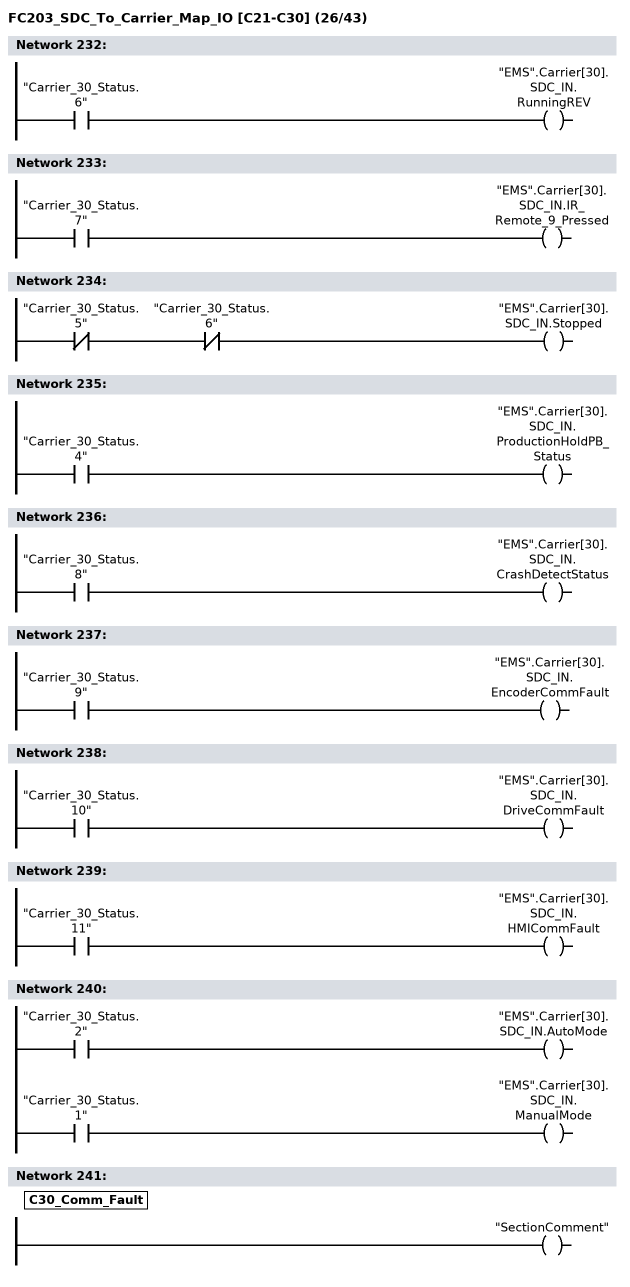
   RUNG wire#powerrail
      Contact( "Carrier_30_Status.6" )
      Coil( "EMS".Carrier[30].SDC_IN.RunningREV )
   END_RUNG
   // the same network as SCL:
   "EMS".Carrier[30].SDC_IN.RunningREV := "Carrier_30_Status.6";
END_REGION

REGION Network 233
   RUNG wire#powerrail
      Contact( "Carrier_30_Status.7" )
      Coil( "EMS".Carrier[30].SDC_IN.IR_Remote_9_Pressed )
   END_RUNG
   // the same network as SCL:
   "EMS".Carrier[30].SDC_IN.IR_Remote_9_Pressed := "Carrier_30_Status.7";
END_REGION

REGION Network 234
   RUNG wire#powerrail
      I_Contact( "Carrier_30_Status.5" )
      I_Contact( "Carrier_30_Status.6" )
      Coil( "EMS".Carrier[30].SDC_IN.Stopped )
   END_RUNG
   // the same network as SCL:
   "EMS".Carrier[30].SDC_IN.Stopped := NOT "Carrier_30_Status.5" AND NOT "Carrier_30_Status.6";
END_REGION

REGION Network 235
   RUNG wire#powerrail
      Contact( "Carrier_30_Status.4" )
      Coil( "EMS".Carrier[30].SDC_IN.ProductionHoldPB_Status )
   END_RUNG
   // the same network as SCL:
   "EMS".Carrier[30].SDC_IN.ProductionHoldPB_Status := "Carrier_30_Status.4";
END_REGION

REGION Network 236
   RUNG wire#powerrail
      Contact( "Carrier_30_Status.8" )
      Coil( "EMS".Carrier[30].SDC_IN.CrashDetectStatus )
   END_RUNG
   // the same network as SCL:
   "EMS".Carrier[30].SDC_IN.CrashDetectStatus := "Carrier_30_Status.8";
END_REGION

REGION Network 237
   RUNG wire#powerrail
      Contact( "Carrier_30_Status.9" )
      Coil( "EMS".Carrier[30].SDC_IN.EncoderCommFault )
   END_RUNG
   // the same network as SCL:
   "EMS".Carrier[30].SDC_IN.EncoderCommFault := "Carrier_30_Status.9";
END_REGION

REGION Network 238
   RUNG wire#powerrail
      Contact( "Carrier_30_Status.10" )
      Coil( "EMS".Carrier[30].SDC_IN.DriveCommFault )
   END_RUNG
   // the same network as SCL:
   "EMS".Carrier[30].SDC_IN.DriveCommFault := "Carrier_30_Status.10";
END_REGION

REGION Network 239
   RUNG wire#powerrail
      Contact( "Carrier_30_Status.11" )
      Coil( "EMS".Carrier[30].SDC_IN.HMICommFault )
   END_RUNG
   // the same network as SCL:
   "EMS".Carrier[30].SDC_IN.HMICommFault := "Carrier_30_Status.11";
END_REGION

REGION Network 240
   RUNG wire#powerrail
      Contact( "Carrier_30_Status.2" )
      Coil( "EMS".Carrier[30].SDC_IN.AutoMode )
   END_RUNG
   RUNG wire#powerrail
      Contact( "Carrier_30_Status.1" )
      Coil( "EMS".Carrier[30].SDC_IN.ManualMode )
   END_RUNG
   // the same network as SCL:
   "EMS".Carrier[30].SDC_IN.AutoMode := "Carrier_30_Status.2";
   "EMS".Carrier[30].SDC_IN.ManualMode := "Carrier_30_Status.1";
END_REGION

REGION Network 241
   Label( C30_Comm_Fault )
   RUNG wire#powerrail
      Coil( "SectionComment" )
   END_RUNG
   // the same network as SCL:
   C30_Comm_Fault:
   "SectionComment" := TRUE;
END_REGION

REGION Network 242
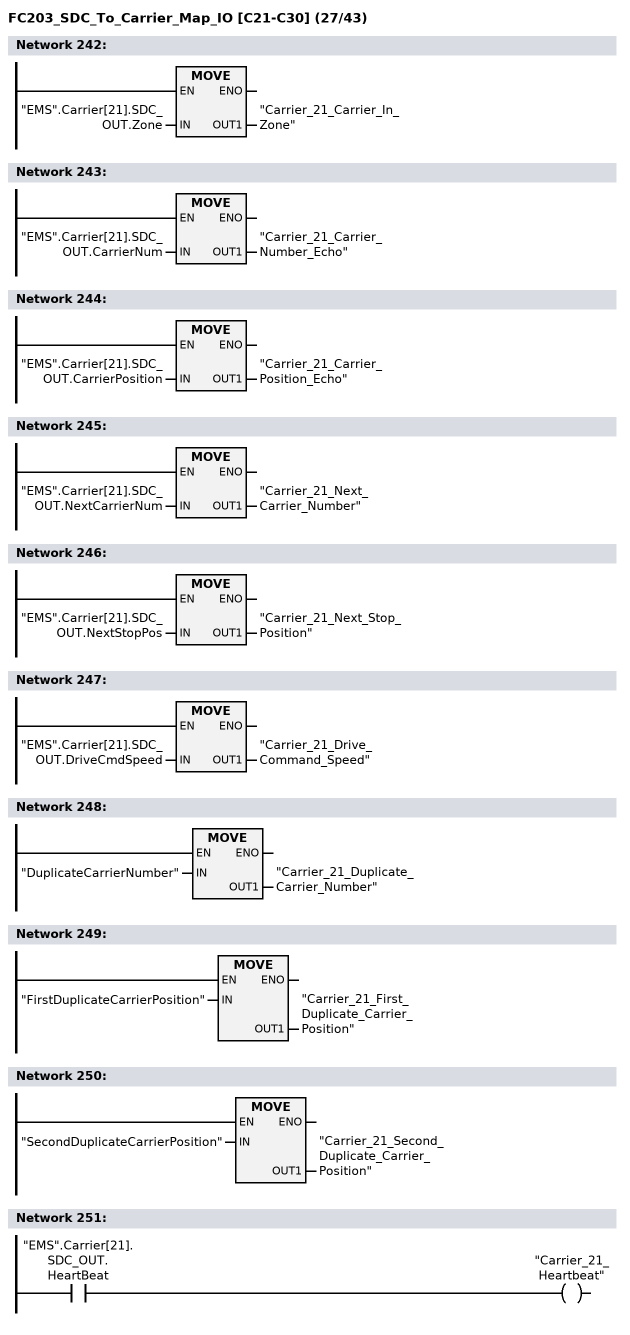
   RUNG wire#powerrail
      Move(in := "EMS".Carrier[21].SDC_OUT.Zone, out1 => "Carrier_21_Carrier_In_Zone")
   END_RUNG
   // the same network as SCL:
   "Carrier_21_Carrier_In_Zone" := "EMS".Carrier[21].SDC_OUT.Zone;
END_REGION

REGION Network 243
   RUNG wire#powerrail
      Move(in := "EMS".Carrier[21].SDC_OUT.CarrierNum, out1 => "Carrier_21_Carrier_Number_Echo")
   END_RUNG
   // the same network as SCL:
   "Carrier_21_Carrier_Number_Echo" := "EMS".Carrier[21].SDC_OUT.CarrierNum;
END_REGION

REGION Network 244
   RUNG wire#powerrail
      Move(in := "EMS".Carrier[21].SDC_OUT.CarrierPosition, out1 => "Carrier_21_Carrier_Position_Echo")
   END_RUNG
   // the same network as SCL:
   "Carrier_21_Carrier_Position_Echo" := "EMS".Carrier[21].SDC_OUT.CarrierPosition;
END_REGION

REGION Network 245
   RUNG wire#powerrail
      Move(in := "EMS".Carrier[21].SDC_OUT.NextCarrierNum, out1 => "Carrier_21_Next_Carrier_Number")
   END_RUNG
   // the same network as SCL:
   "Carrier_21_Next_Carrier_Number" := "EMS".Carrier[21].SDC_OUT.NextCarrierNum;
END_REGION

REGION Network 246
   RUNG wire#powerrail
      Move(in := "EMS".Carrier[21].SDC_OUT.NextStopPos, out1 => "Carrier_21_Next_Stop_Position")
   END_RUNG
   // the same network as SCL:
   "Carrier_21_Next_Stop_Position" := "EMS".Carrier[21].SDC_OUT.NextStopPos;
END_REGION

REGION Network 247
   RUNG wire#powerrail
      Move(in := "EMS".Carrier[21].SDC_OUT.DriveCmdSpeed, out1 => "Carrier_21_Drive_Command_Speed")
   END_RUNG
   // the same network as SCL:
   "Carrier_21_Drive_Command_Speed" := "EMS".Carrier[21].SDC_OUT.DriveCmdSpeed;
END_REGION

REGION Network 248
   RUNG wire#powerrail
      Move(in := "DuplicateCarrierNumber", out1 => "Carrier_21_Duplicate_Carrier_Number")
   END_RUNG
   // the same network as SCL:
   "Carrier_21_Duplicate_Carrier_Number" := "DuplicateCarrierNumber";
END_REGION

REGION Network 249
   RUNG wire#powerrail
      Move(in := "FirstDuplicateCarrierPosition", out1 => "Carrier_21_First_Duplicate_Carrier_Position")
   END_RUNG
   // the same network as SCL:
   "Carrier_21_First_Duplicate_Carrier_Position" := "FirstDuplicateCarrierPosition";
END_REGION

REGION Network 250
   RUNG wire#powerrail
      Move(in := "SecondDuplicateCarrierPosition", out1 => "Carrier_21_Second_Duplicate_Carrier_Position")
   END_RUNG
   // the same network as SCL:
   "Carrier_21_Second_Duplicate_Carrier_Position" := "SecondDuplicateCarrierPosition";
END_REGION

REGION Network 251
   RUNG wire#powerrail
      Contact( "EMS".Carrier[21].SDC_OUT.HeartBeat )
      Coil( "Carrier_21_Heartbeat" )
   END_RUNG
   // the same network as SCL:
   "Carrier_21_Heartbeat" := "EMS".Carrier[21].SDC_OUT.HeartBeat;
END_REGION

REGION Network 252
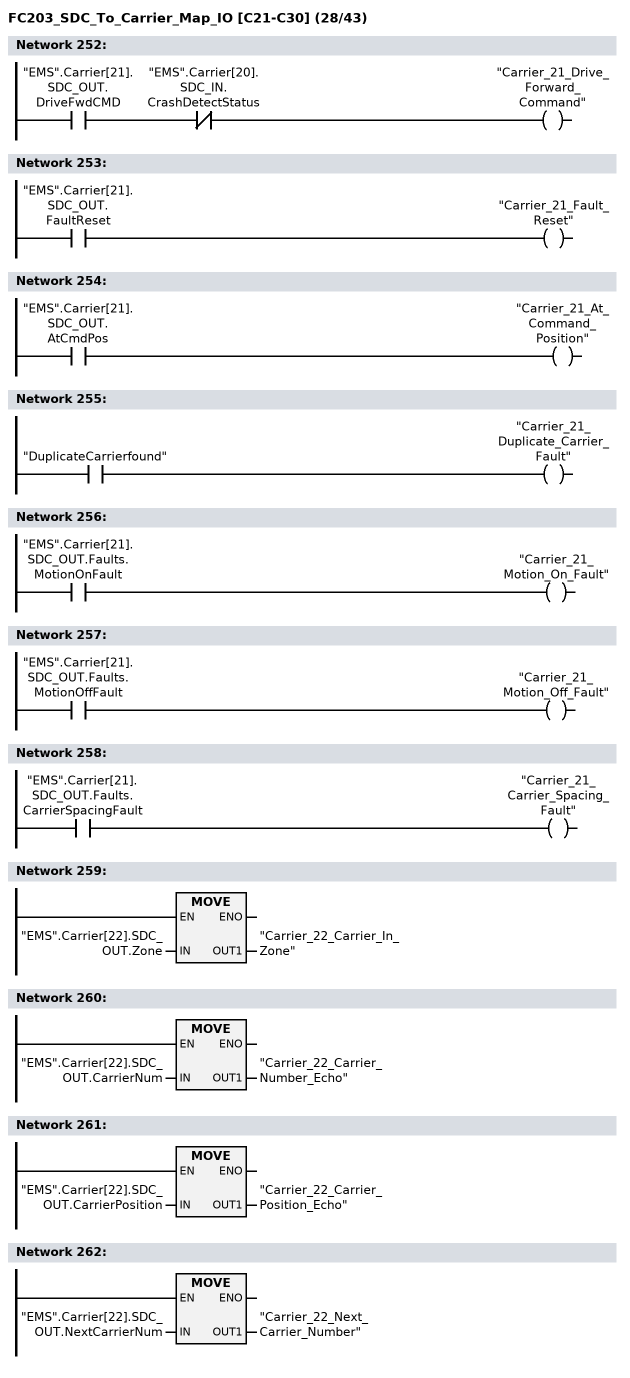
   RUNG wire#powerrail
      Contact( "EMS".Carrier[21].SDC_OUT.DriveFwdCMD )
      I_Contact( "EMS".Carrier[20].SDC_IN.CrashDetectStatus )
      Coil( "Carrier_21_Drive_Forward_Command" )
   END_RUNG
   // the same network as SCL:
   "Carrier_21_Drive_Forward_Command" := "EMS".Carrier[21].SDC_OUT.DriveFwdCMD AND NOT "EMS".Carrier[20].SDC_IN.CrashDetectStatus;
END_REGION

REGION Network 253
   RUNG wire#powerrail
      Contact( "EMS".Carrier[21].SDC_OUT.FaultReset )
      Coil( "Carrier_21_Fault_Reset" )
   END_RUNG
   // the same network as SCL:
   "Carrier_21_Fault_Reset" := "EMS".Carrier[21].SDC_OUT.FaultReset;
END_REGION

REGION Network 254
   RUNG wire#powerrail
      Contact( "EMS".Carrier[21].SDC_OUT.AtCmdPos )
      Coil( "Carrier_21_At_Command_Position" )
   END_RUNG
   // the same network as SCL:
   "Carrier_21_At_Command_Position" := "EMS".Carrier[21].SDC_OUT.AtCmdPos;
END_REGION

REGION Network 255
   RUNG wire#powerrail
      Contact( "DuplicateCarrierfound" )
      Coil( "Carrier_21_Duplicate_Carrier_Fault" )
   END_RUNG
   // the same network as SCL:
   "Carrier_21_Duplicate_Carrier_Fault" := "DuplicateCarrierfound";
END_REGION

REGION Network 256
   RUNG wire#powerrail
      Contact( "EMS".Carrier[21].SDC_OUT.Faults.MotionOnFault )
      Coil( "Carrier_21_Motion_On_Fault" )
   END_RUNG
   // the same network as SCL:
   "Carrier_21_Motion_On_Fault" := "EMS".Carrier[21].SDC_OUT.Faults.MotionOnFault;
END_REGION

REGION Network 257
   RUNG wire#powerrail
      Contact( "EMS".Carrier[21].SDC_OUT.Faults.MotionOffFault )
      Coil( "Carrier_21_Motion_Off_Fault" )
   END_RUNG
   // the same network as SCL:
   "Carrier_21_Motion_Off_Fault" := "EMS".Carrier[21].SDC_OUT.Faults.MotionOffFault;
END_REGION

REGION Network 258
   RUNG wire#powerrail
      Contact( "EMS".Carrier[21].SDC_OUT.Faults.CarrierSpacingFault )
      Coil( "Carrier_21_Carrier_Spacing_Fault" )
   END_RUNG
   // the same network as SCL:
   "Carrier_21_Carrier_Spacing_Fault" := "EMS".Carrier[21].SDC_OUT.Faults.CarrierSpacingFault;
END_REGION

REGION Network 259
   RUNG wire#powerrail
      Move(in := "EMS".Carrier[22].SDC_OUT.Zone, out1 => "Carrier_22_Carrier_In_Zone")
   END_RUNG
   // the same network as SCL:
   "Carrier_22_Carrier_In_Zone" := "EMS".Carrier[22].SDC_OUT.Zone;
END_REGION

REGION Network 260
   RUNG wire#powerrail
      Move(in := "EMS".Carrier[22].SDC_OUT.CarrierNum, out1 => "Carrier_22_Carrier_Number_Echo")
   END_RUNG
   // the same network as SCL:
   "Carrier_22_Carrier_Number_Echo" := "EMS".Carrier[22].SDC_OUT.CarrierNum;
END_REGION

REGION Network 261
   RUNG wire#powerrail
      Move(in := "EMS".Carrier[22].SDC_OUT.CarrierPosition, out1 => "Carrier_22_Carrier_Position_Echo")
   END_RUNG
   // the same network as SCL:
   "Carrier_22_Carrier_Position_Echo" := "EMS".Carrier[22].SDC_OUT.CarrierPosition;
END_REGION

REGION Network 262
   RUNG wire#powerrail
      Move(in := "EMS".Carrier[22].SDC_OUT.NextCarrierNum, out1 => "Carrier_22_Next_Carrier_Number")
   END_RUNG
   // the same network as SCL:
   "Carrier_22_Next_Carrier_Number" := "EMS".Carrier[22].SDC_OUT.NextCarrierNum;
END_REGION

REGION Network 263
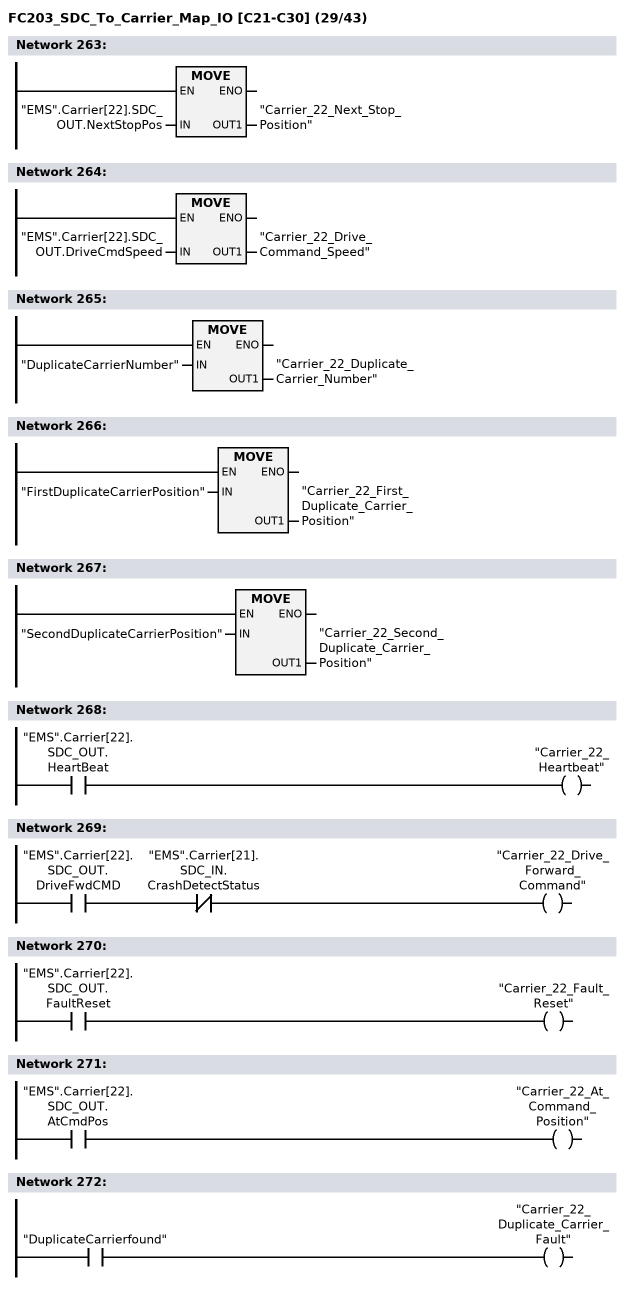
   RUNG wire#powerrail
      Move(in := "EMS".Carrier[22].SDC_OUT.NextStopPos, out1 => "Carrier_22_Next_Stop_Position")
   END_RUNG
   // the same network as SCL:
   "Carrier_22_Next_Stop_Position" := "EMS".Carrier[22].SDC_OUT.NextStopPos;
END_REGION

REGION Network 264
   RUNG wire#powerrail
      Move(in := "EMS".Carrier[22].SDC_OUT.DriveCmdSpeed, out1 => "Carrier_22_Drive_Command_Speed")
   END_RUNG
   // the same network as SCL:
   "Carrier_22_Drive_Command_Speed" := "EMS".Carrier[22].SDC_OUT.DriveCmdSpeed;
END_REGION

REGION Network 265
   RUNG wire#powerrail
      Move(in := "DuplicateCarrierNumber", out1 => "Carrier_22_Duplicate_Carrier_Number")
   END_RUNG
   // the same network as SCL:
   "Carrier_22_Duplicate_Carrier_Number" := "DuplicateCarrierNumber";
END_REGION

REGION Network 266
   RUNG wire#powerrail
      Move(in := "FirstDuplicateCarrierPosition", out1 => "Carrier_22_First_Duplicate_Carrier_Position")
   END_RUNG
   // the same network as SCL:
   "Carrier_22_First_Duplicate_Carrier_Position" := "FirstDuplicateCarrierPosition";
END_REGION

REGION Network 267
   RUNG wire#powerrail
      Move(in := "SecondDuplicateCarrierPosition", out1 => "Carrier_22_Second_Duplicate_Carrier_Position")
   END_RUNG
   // the same network as SCL:
   "Carrier_22_Second_Duplicate_Carrier_Position" := "SecondDuplicateCarrierPosition";
END_REGION

REGION Network 268
   RUNG wire#powerrail
      Contact( "EMS".Carrier[22].SDC_OUT.HeartBeat )
      Coil( "Carrier_22_Heartbeat" )
   END_RUNG
   // the same network as SCL:
   "Carrier_22_Heartbeat" := "EMS".Carrier[22].SDC_OUT.HeartBeat;
END_REGION

REGION Network 269
   RUNG wire#powerrail
      Contact( "EMS".Carrier[22].SDC_OUT.DriveFwdCMD )
      I_Contact( "EMS".Carrier[21].SDC_IN.CrashDetectStatus )
      Coil( "Carrier_22_Drive_Forward_Command" )
   END_RUNG
   // the same network as SCL:
   "Carrier_22_Drive_Forward_Command" := "EMS".Carrier[22].SDC_OUT.DriveFwdCMD AND NOT "EMS".Carrier[21].SDC_IN.CrashDetectStatus;
END_REGION

REGION Network 270
   RUNG wire#powerrail
      Contact( "EMS".Carrier[22].SDC_OUT.FaultReset )
      Coil( "Carrier_22_Fault_Reset" )
   END_RUNG
   // the same network as SCL:
   "Carrier_22_Fault_Reset" := "EMS".Carrier[22].SDC_OUT.FaultReset;
END_REGION

REGION Network 271
   RUNG wire#powerrail
      Contact( "EMS".Carrier[22].SDC_OUT.AtCmdPos )
      Coil( "Carrier_22_At_Command_Position" )
   END_RUNG
   // the same network as SCL:
   "Carrier_22_At_Command_Position" := "EMS".Carrier[22].SDC_OUT.AtCmdPos;
END_REGION

REGION Network 272
   RUNG wire#powerrail
      Contact( "DuplicateCarrierfound" )
      Coil( "Carrier_22_Duplicate_Carrier_Fault" )
   END_RUNG
   // the same network as SCL:
   "Carrier_22_Duplicate_Carrier_Fault" := "DuplicateCarrierfound";
END_REGION

REGION Network 273
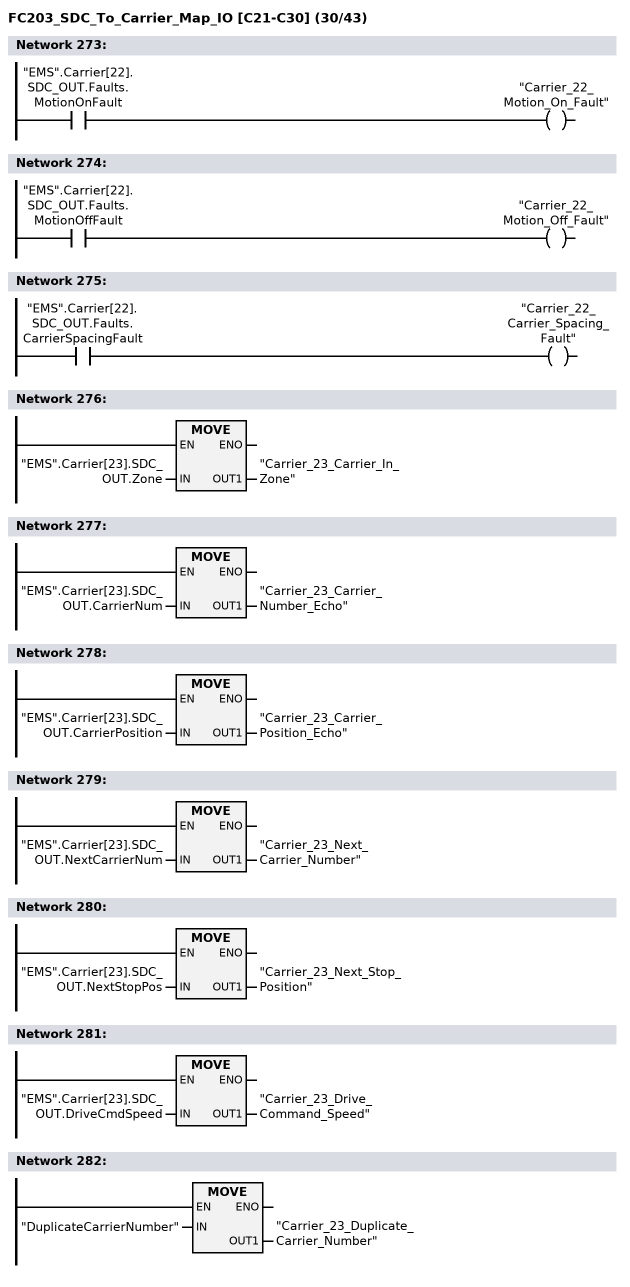
   RUNG wire#powerrail
      Contact( "EMS".Carrier[22].SDC_OUT.Faults.MotionOnFault )
      Coil( "Carrier_22_Motion_On_Fault" )
   END_RUNG
   // the same network as SCL:
   "Carrier_22_Motion_On_Fault" := "EMS".Carrier[22].SDC_OUT.Faults.MotionOnFault;
END_REGION

REGION Network 274
   RUNG wire#powerrail
      Contact( "EMS".Carrier[22].SDC_OUT.Faults.MotionOffFault )
      Coil( "Carrier_22_Motion_Off_Fault" )
   END_RUNG
   // the same network as SCL:
   "Carrier_22_Motion_Off_Fault" := "EMS".Carrier[22].SDC_OUT.Faults.MotionOffFault;
END_REGION

REGION Network 275
   RUNG wire#powerrail
      Contact( "EMS".Carrier[22].SDC_OUT.Faults.CarrierSpacingFault )
      Coil( "Carrier_22_Carrier_Spacing_Fault" )
   END_RUNG
   // the same network as SCL:
   "Carrier_22_Carrier_Spacing_Fault" := "EMS".Carrier[22].SDC_OUT.Faults.CarrierSpacingFault;
END_REGION

REGION Network 276
   RUNG wire#powerrail
      Move(in := "EMS".Carrier[23].SDC_OUT.Zone, out1 => "Carrier_23_Carrier_In_Zone")
   END_RUNG
   // the same network as SCL:
   "Carrier_23_Carrier_In_Zone" := "EMS".Carrier[23].SDC_OUT.Zone;
END_REGION

REGION Network 277
   RUNG wire#powerrail
      Move(in := "EMS".Carrier[23].SDC_OUT.CarrierNum, out1 => "Carrier_23_Carrier_Number_Echo")
   END_RUNG
   // the same network as SCL:
   "Carrier_23_Carrier_Number_Echo" := "EMS".Carrier[23].SDC_OUT.CarrierNum;
END_REGION

REGION Network 278
   RUNG wire#powerrail
      Move(in := "EMS".Carrier[23].SDC_OUT.CarrierPosition, out1 => "Carrier_23_Carrier_Position_Echo")
   END_RUNG
   // the same network as SCL:
   "Carrier_23_Carrier_Position_Echo" := "EMS".Carrier[23].SDC_OUT.CarrierPosition;
END_REGION

REGION Network 279
   RUNG wire#powerrail
      Move(in := "EMS".Carrier[23].SDC_OUT.NextCarrierNum, out1 => "Carrier_23_Next_Carrier_Number")
   END_RUNG
   // the same network as SCL:
   "Carrier_23_Next_Carrier_Number" := "EMS".Carrier[23].SDC_OUT.NextCarrierNum;
END_REGION

REGION Network 280
   RUNG wire#powerrail
      Move(in := "EMS".Carrier[23].SDC_OUT.NextStopPos, out1 => "Carrier_23_Next_Stop_Position")
   END_RUNG
   // the same network as SCL:
   "Carrier_23_Next_Stop_Position" := "EMS".Carrier[23].SDC_OUT.NextStopPos;
END_REGION

REGION Network 281
   RUNG wire#powerrail
      Move(in := "EMS".Carrier[23].SDC_OUT.DriveCmdSpeed, out1 => "Carrier_23_Drive_Command_Speed")
   END_RUNG
   // the same network as SCL:
   "Carrier_23_Drive_Command_Speed" := "EMS".Carrier[23].SDC_OUT.DriveCmdSpeed;
END_REGION

REGION Network 282
   RUNG wire#powerrail
      Move(in := "DuplicateCarrierNumber", out1 => "Carrier_23_Duplicate_Carrier_Number")
   END_RUNG
   // the same network as SCL:
   "Carrier_23_Duplicate_Carrier_Number" := "DuplicateCarrierNumber";
END_REGION

REGION Network 283
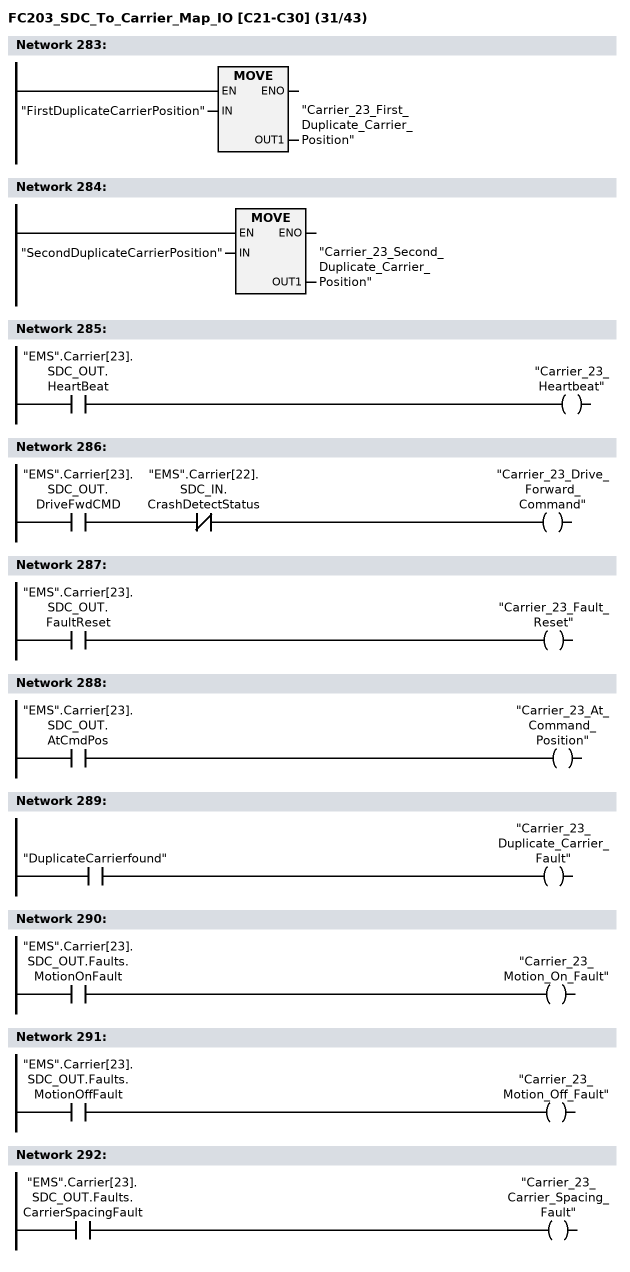
   RUNG wire#powerrail
      Move(in := "FirstDuplicateCarrierPosition", out1 => "Carrier_23_First_Duplicate_Carrier_Position")
   END_RUNG
   // the same network as SCL:
   "Carrier_23_First_Duplicate_Carrier_Position" := "FirstDuplicateCarrierPosition";
END_REGION

REGION Network 284
   RUNG wire#powerrail
      Move(in := "SecondDuplicateCarrierPosition", out1 => "Carrier_23_Second_Duplicate_Carrier_Position")
   END_RUNG
   // the same network as SCL:
   "Carrier_23_Second_Duplicate_Carrier_Position" := "SecondDuplicateCarrierPosition";
END_REGION

REGION Network 285
   RUNG wire#powerrail
      Contact( "EMS".Carrier[23].SDC_OUT.HeartBeat )
      Coil( "Carrier_23_Heartbeat" )
   END_RUNG
   // the same network as SCL:
   "Carrier_23_Heartbeat" := "EMS".Carrier[23].SDC_OUT.HeartBeat;
END_REGION

REGION Network 286
   RUNG wire#powerrail
      Contact( "EMS".Carrier[23].SDC_OUT.DriveFwdCMD )
      I_Contact( "EMS".Carrier[22].SDC_IN.CrashDetectStatus )
      Coil( "Carrier_23_Drive_Forward_Command" )
   END_RUNG
   // the same network as SCL:
   "Carrier_23_Drive_Forward_Command" := "EMS".Carrier[23].SDC_OUT.DriveFwdCMD AND NOT "EMS".Carrier[22].SDC_IN.CrashDetectStatus;
END_REGION

REGION Network 287
   RUNG wire#powerrail
      Contact( "EMS".Carrier[23].SDC_OUT.FaultReset )
      Coil( "Carrier_23_Fault_Reset" )
   END_RUNG
   // the same network as SCL:
   "Carrier_23_Fault_Reset" := "EMS".Carrier[23].SDC_OUT.FaultReset;
END_REGION

REGION Network 288
   RUNG wire#powerrail
      Contact( "EMS".Carrier[23].SDC_OUT.AtCmdPos )
      Coil( "Carrier_23_At_Command_Position" )
   END_RUNG
   // the same network as SCL:
   "Carrier_23_At_Command_Position" := "EMS".Carrier[23].SDC_OUT.AtCmdPos;
END_REGION

REGION Network 289
   RUNG wire#powerrail
      Contact( "DuplicateCarrierfound" )
      Coil( "Carrier_23_Duplicate_Carrier_Fault" )
   END_RUNG
   // the same network as SCL:
   "Carrier_23_Duplicate_Carrier_Fault" := "DuplicateCarrierfound";
END_REGION

REGION Network 290
   RUNG wire#powerrail
      Contact( "EMS".Carrier[23].SDC_OUT.Faults.MotionOnFault )
      Coil( "Carrier_23_Motion_On_Fault" )
   END_RUNG
   // the same network as SCL:
   "Carrier_23_Motion_On_Fault" := "EMS".Carrier[23].SDC_OUT.Faults.MotionOnFault;
END_REGION

REGION Network 291
   RUNG wire#powerrail
      Contact( "EMS".Carrier[23].SDC_OUT.Faults.MotionOffFault )
      Coil( "Carrier_23_Motion_Off_Fault" )
   END_RUNG
   // the same network as SCL:
   "Carrier_23_Motion_Off_Fault" := "EMS".Carrier[23].SDC_OUT.Faults.MotionOffFault;
END_REGION

REGION Network 292
   RUNG wire#powerrail
      Contact( "EMS".Carrier[23].SDC_OUT.Faults.CarrierSpacingFault )
      Coil( "Carrier_23_Carrier_Spacing_Fault" )
   END_RUNG
   // the same network as SCL:
   "Carrier_23_Carrier_Spacing_Fault" := "EMS".Carrier[23].SDC_OUT.Faults.CarrierSpacingFault;
END_REGION

REGION Network 293
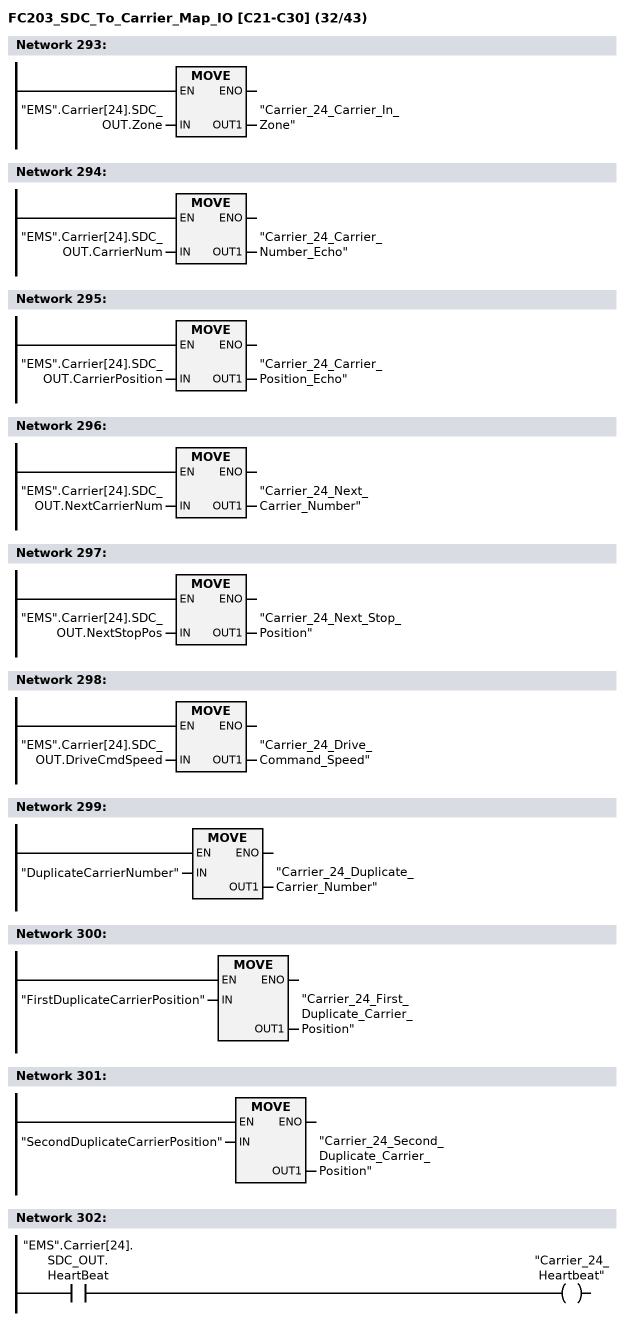
   RUNG wire#powerrail
      Move(in := "EMS".Carrier[24].SDC_OUT.Zone, out1 => "Carrier_24_Carrier_In_Zone")
   END_RUNG
   // the same network as SCL:
   "Carrier_24_Carrier_In_Zone" := "EMS".Carrier[24].SDC_OUT.Zone;
END_REGION

REGION Network 294
   RUNG wire#powerrail
      Move(in := "EMS".Carrier[24].SDC_OUT.CarrierNum, out1 => "Carrier_24_Carrier_Number_Echo")
   END_RUNG
   // the same network as SCL:
   "Carrier_24_Carrier_Number_Echo" := "EMS".Carrier[24].SDC_OUT.CarrierNum;
END_REGION

REGION Network 295
   RUNG wire#powerrail
      Move(in := "EMS".Carrier[24].SDC_OUT.CarrierPosition, out1 => "Carrier_24_Carrier_Position_Echo")
   END_RUNG
   // the same network as SCL:
   "Carrier_24_Carrier_Position_Echo" := "EMS".Carrier[24].SDC_OUT.CarrierPosition;
END_REGION

REGION Network 296
   RUNG wire#powerrail
      Move(in := "EMS".Carrier[24].SDC_OUT.NextCarrierNum, out1 => "Carrier_24_Next_Carrier_Number")
   END_RUNG
   // the same network as SCL:
   "Carrier_24_Next_Carrier_Number" := "EMS".Carrier[24].SDC_OUT.NextCarrierNum;
END_REGION

REGION Network 297
   RUNG wire#powerrail
      Move(in := "EMS".Carrier[24].SDC_OUT.NextStopPos, out1 => "Carrier_24_Next_Stop_Position")
   END_RUNG
   // the same network as SCL:
   "Carrier_24_Next_Stop_Position" := "EMS".Carrier[24].SDC_OUT.NextStopPos;
END_REGION

REGION Network 298
   RUNG wire#powerrail
      Move(in := "EMS".Carrier[24].SDC_OUT.DriveCmdSpeed, out1 => "Carrier_24_Drive_Command_Speed")
   END_RUNG
   // the same network as SCL:
   "Carrier_24_Drive_Command_Speed" := "EMS".Carrier[24].SDC_OUT.DriveCmdSpeed;
END_REGION

REGION Network 299
   RUNG wire#powerrail
      Move(in := "DuplicateCarrierNumber", out1 => "Carrier_24_Duplicate_Carrier_Number")
   END_RUNG
   // the same network as SCL:
   "Carrier_24_Duplicate_Carrier_Number" := "DuplicateCarrierNumber";
END_REGION

REGION Network 300
   RUNG wire#powerrail
      Move(in := "FirstDuplicateCarrierPosition", out1 => "Carrier_24_First_Duplicate_Carrier_Position")
   END_RUNG
   // the same network as SCL:
   "Carrier_24_First_Duplicate_Carrier_Position" := "FirstDuplicateCarrierPosition";
END_REGION

REGION Network 301
   RUNG wire#powerrail
      Move(in := "SecondDuplicateCarrierPosition", out1 => "Carrier_24_Second_Duplicate_Carrier_Position")
   END_RUNG
   // the same network as SCL:
   "Carrier_24_Second_Duplicate_Carrier_Position" := "SecondDuplicateCarrierPosition";
END_REGION

REGION Network 302
   RUNG wire#powerrail
      Contact( "EMS".Carrier[24].SDC_OUT.HeartBeat )
      Coil( "Carrier_24_Heartbeat" )
   END_RUNG
   // the same network as SCL:
   "Carrier_24_Heartbeat" := "EMS".Carrier[24].SDC_OUT.HeartBeat;
END_REGION

REGION Network 303
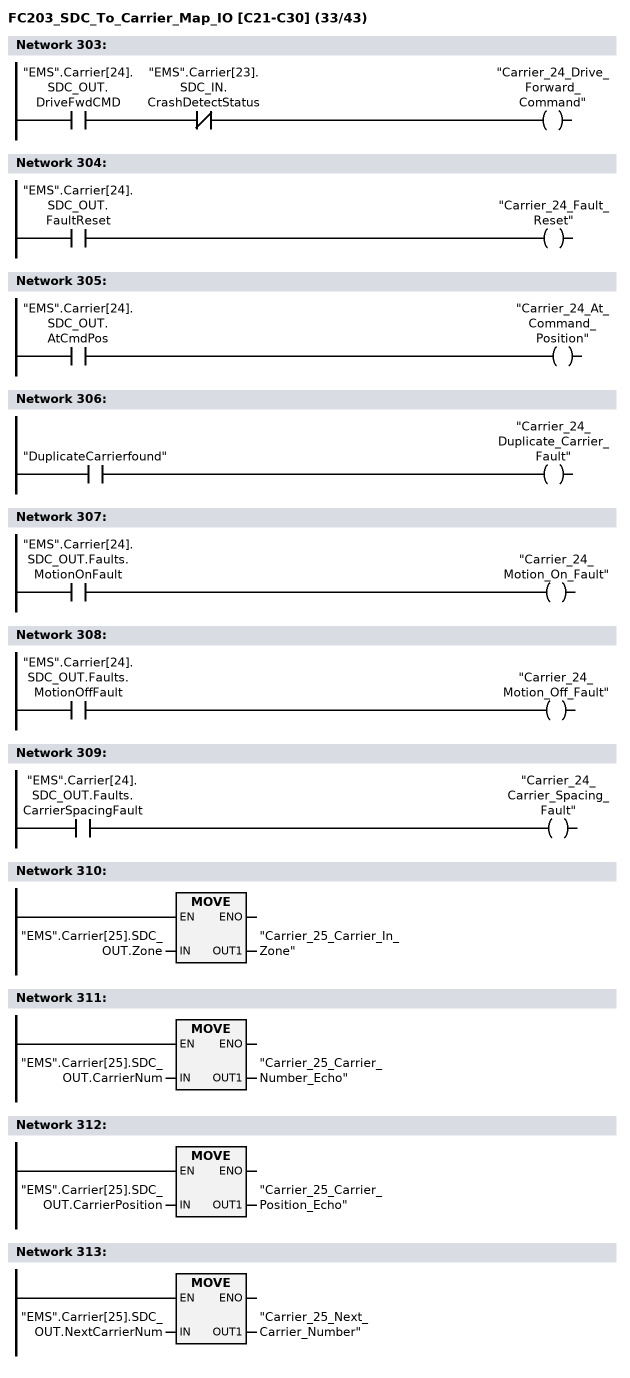
   RUNG wire#powerrail
      Contact( "EMS".Carrier[24].SDC_OUT.DriveFwdCMD )
      I_Contact( "EMS".Carrier[23].SDC_IN.CrashDetectStatus )
      Coil( "Carrier_24_Drive_Forward_Command" )
   END_RUNG
   // the same network as SCL:
   "Carrier_24_Drive_Forward_Command" := "EMS".Carrier[24].SDC_OUT.DriveFwdCMD AND NOT "EMS".Carrier[23].SDC_IN.CrashDetectStatus;
END_REGION

REGION Network 304
   RUNG wire#powerrail
      Contact( "EMS".Carrier[24].SDC_OUT.FaultReset )
      Coil( "Carrier_24_Fault_Reset" )
   END_RUNG
   // the same network as SCL:
   "Carrier_24_Fault_Reset" := "EMS".Carrier[24].SDC_OUT.FaultReset;
END_REGION

REGION Network 305
   RUNG wire#powerrail
      Contact( "EMS".Carrier[24].SDC_OUT.AtCmdPos )
      Coil( "Carrier_24_At_Command_Position" )
   END_RUNG
   // the same network as SCL:
   "Carrier_24_At_Command_Position" := "EMS".Carrier[24].SDC_OUT.AtCmdPos;
END_REGION

REGION Network 306
   RUNG wire#powerrail
      Contact( "DuplicateCarrierfound" )
      Coil( "Carrier_24_Duplicate_Carrier_Fault" )
   END_RUNG
   // the same network as SCL:
   "Carrier_24_Duplicate_Carrier_Fault" := "DuplicateCarrierfound";
END_REGION

REGION Network 307
   RUNG wire#powerrail
      Contact( "EMS".Carrier[24].SDC_OUT.Faults.MotionOnFault )
      Coil( "Carrier_24_Motion_On_Fault" )
   END_RUNG
   // the same network as SCL:
   "Carrier_24_Motion_On_Fault" := "EMS".Carrier[24].SDC_OUT.Faults.MotionOnFault;
END_REGION

REGION Network 308
   RUNG wire#powerrail
      Contact( "EMS".Carrier[24].SDC_OUT.Faults.MotionOffFault )
      Coil( "Carrier_24_Motion_Off_Fault" )
   END_RUNG
   // the same network as SCL:
   "Carrier_24_Motion_Off_Fault" := "EMS".Carrier[24].SDC_OUT.Faults.MotionOffFault;
END_REGION

REGION Network 309
   RUNG wire#powerrail
      Contact( "EMS".Carrier[24].SDC_OUT.Faults.CarrierSpacingFault )
      Coil( "Carrier_24_Carrier_Spacing_Fault" )
   END_RUNG
   // the same network as SCL:
   "Carrier_24_Carrier_Spacing_Fault" := "EMS".Carrier[24].SDC_OUT.Faults.CarrierSpacingFault;
END_REGION

REGION Network 310
   RUNG wire#powerrail
      Move(in := "EMS".Carrier[25].SDC_OUT.Zone, out1 => "Carrier_25_Carrier_In_Zone")
   END_RUNG
   // the same network as SCL:
   "Carrier_25_Carrier_In_Zone" := "EMS".Carrier[25].SDC_OUT.Zone;
END_REGION

REGION Network 311
   RUNG wire#powerrail
      Move(in := "EMS".Carrier[25].SDC_OUT.CarrierNum, out1 => "Carrier_25_Carrier_Number_Echo")
   END_RUNG
   // the same network as SCL:
   "Carrier_25_Carrier_Number_Echo" := "EMS".Carrier[25].SDC_OUT.CarrierNum;
END_REGION

REGION Network 312
   RUNG wire#powerrail
      Move(in := "EMS".Carrier[25].SDC_OUT.CarrierPosition, out1 => "Carrier_25_Carrier_Position_Echo")
   END_RUNG
   // the same network as SCL:
   "Carrier_25_Carrier_Position_Echo" := "EMS".Carrier[25].SDC_OUT.CarrierPosition;
END_REGION

REGION Network 313
   RUNG wire#powerrail
      Move(in := "EMS".Carrier[25].SDC_OUT.NextCarrierNum, out1 => "Carrier_25_Next_Carrier_Number")
   END_RUNG
   // the same network as SCL:
   "Carrier_25_Next_Carrier_Number" := "EMS".Carrier[25].SDC_OUT.NextCarrierNum;
END_REGION

REGION Network 314
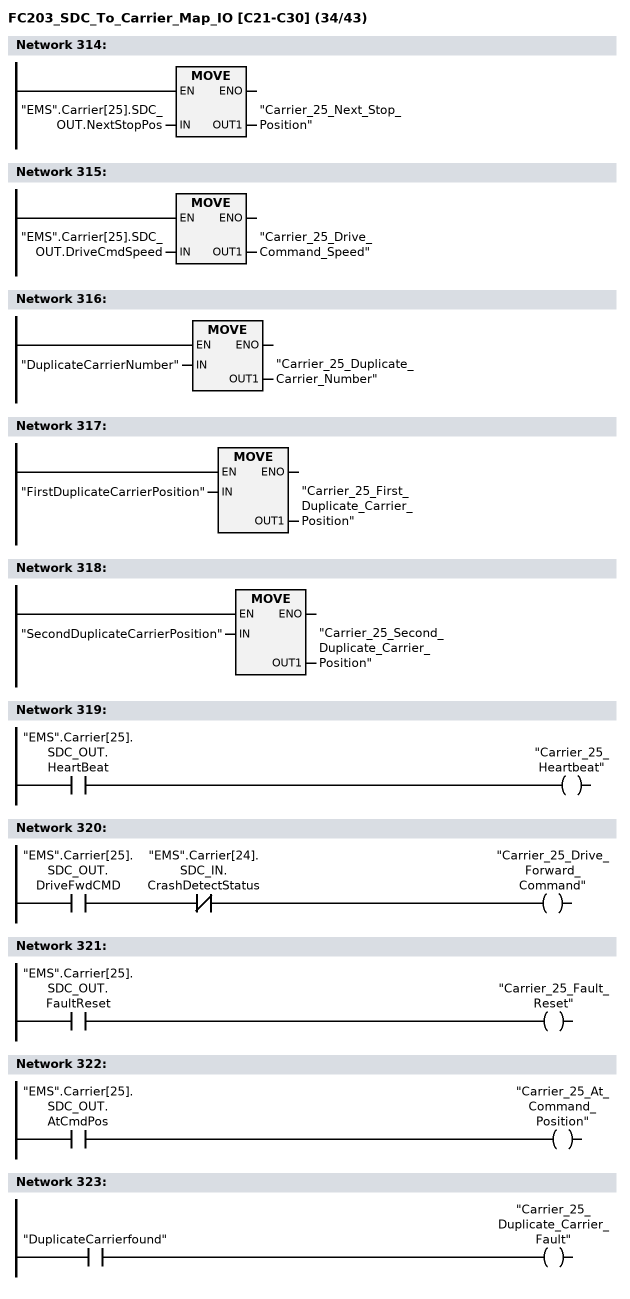
   RUNG wire#powerrail
      Move(in := "EMS".Carrier[25].SDC_OUT.NextStopPos, out1 => "Carrier_25_Next_Stop_Position")
   END_RUNG
   // the same network as SCL:
   "Carrier_25_Next_Stop_Position" := "EMS".Carrier[25].SDC_OUT.NextStopPos;
END_REGION

REGION Network 315
   RUNG wire#powerrail
      Move(in := "EMS".Carrier[25].SDC_OUT.DriveCmdSpeed, out1 => "Carrier_25_Drive_Command_Speed")
   END_RUNG
   // the same network as SCL:
   "Carrier_25_Drive_Command_Speed" := "EMS".Carrier[25].SDC_OUT.DriveCmdSpeed;
END_REGION

REGION Network 316
   RUNG wire#powerrail
      Move(in := "DuplicateCarrierNumber", out1 => "Carrier_25_Duplicate_Carrier_Number")
   END_RUNG
   // the same network as SCL:
   "Carrier_25_Duplicate_Carrier_Number" := "DuplicateCarrierNumber";
END_REGION

REGION Network 317
   RUNG wire#powerrail
      Move(in := "FirstDuplicateCarrierPosition", out1 => "Carrier_25_First_Duplicate_Carrier_Position")
   END_RUNG
   // the same network as SCL:
   "Carrier_25_First_Duplicate_Carrier_Position" := "FirstDuplicateCarrierPosition";
END_REGION

REGION Network 318
   RUNG wire#powerrail
      Move(in := "SecondDuplicateCarrierPosition", out1 => "Carrier_25_Second_Duplicate_Carrier_Position")
   END_RUNG
   // the same network as SCL:
   "Carrier_25_Second_Duplicate_Carrier_Position" := "SecondDuplicateCarrierPosition";
END_REGION

REGION Network 319
   RUNG wire#powerrail
      Contact( "EMS".Carrier[25].SDC_OUT.HeartBeat )
      Coil( "Carrier_25_Heartbeat" )
   END_RUNG
   // the same network as SCL:
   "Carrier_25_Heartbeat" := "EMS".Carrier[25].SDC_OUT.HeartBeat;
END_REGION

REGION Network 320
   RUNG wire#powerrail
      Contact( "EMS".Carrier[25].SDC_OUT.DriveFwdCMD )
      I_Contact( "EMS".Carrier[24].SDC_IN.CrashDetectStatus )
      Coil( "Carrier_25_Drive_Forward_Command" )
   END_RUNG
   // the same network as SCL:
   "Carrier_25_Drive_Forward_Command" := "EMS".Carrier[25].SDC_OUT.DriveFwdCMD AND NOT "EMS".Carrier[24].SDC_IN.CrashDetectStatus;
END_REGION

REGION Network 321
   RUNG wire#powerrail
      Contact( "EMS".Carrier[25].SDC_OUT.FaultReset )
      Coil( "Carrier_25_Fault_Reset" )
   END_RUNG
   // the same network as SCL:
   "Carrier_25_Fault_Reset" := "EMS".Carrier[25].SDC_OUT.FaultReset;
END_REGION

REGION Network 322
   RUNG wire#powerrail
      Contact( "EMS".Carrier[25].SDC_OUT.AtCmdPos )
      Coil( "Carrier_25_At_Command_Position" )
   END_RUNG
   // the same network as SCL:
   "Carrier_25_At_Command_Position" := "EMS".Carrier[25].SDC_OUT.AtCmdPos;
END_REGION

REGION Network 323
   RUNG wire#powerrail
      Contact( "DuplicateCarrierfound" )
      Coil( "Carrier_25_Duplicate_Carrier_Fault" )
   END_RUNG
   // the same network as SCL:
   "Carrier_25_Duplicate_Carrier_Fault" := "DuplicateCarrierfound";
END_REGION

REGION Network 324
